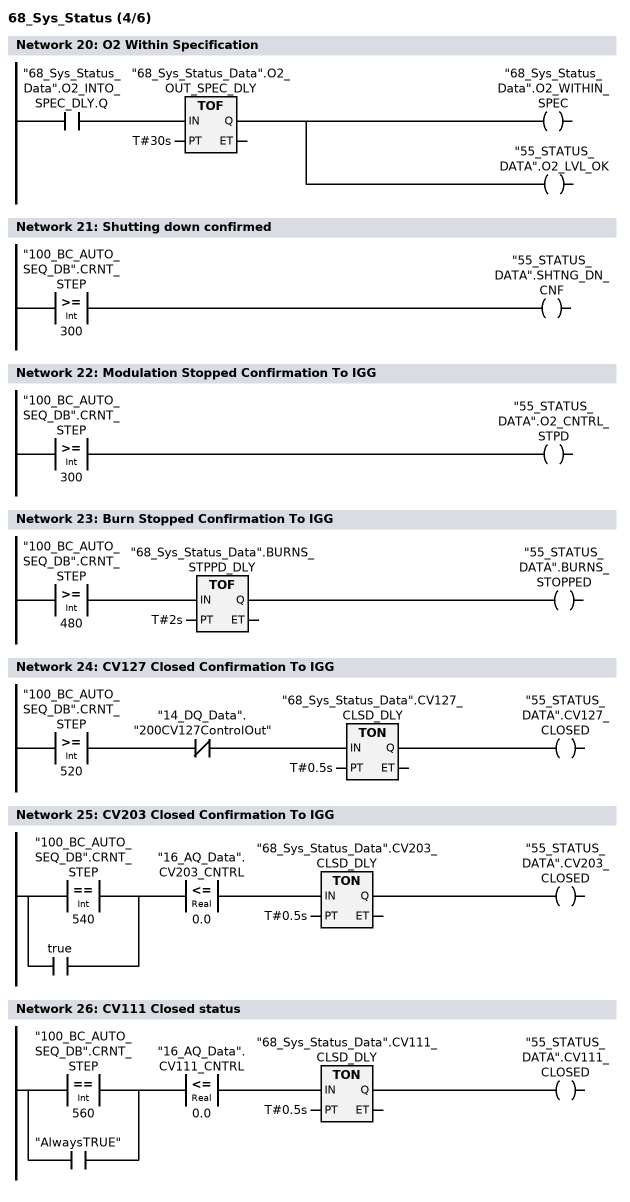
   "68_Sys_Status_Data".O2_OUT_SPEC_DLY.TOF(IN := "68_Sys_Status_Data".O2_INTO_SPEC_DLY.Q, PT := T#30s);
   "68_Sys_Status_Data".O2_WITHIN_SPEC := "68_Sys_Status_Data".O2_OUT_SPEC_DLY.Q;
   "55_STATUS_DATA".O2_LVL_OK := "68_Sys_Status_Data".O2_OUT_SPEC_DLY.Q;
END_REGION

REGION Network 21: Shutting down confirmed
   RUNG wire#powerrail
      { S7_Templates := "SrcType := Int" } GE_Contact(in1 := "100_BC_AUTO_SEQ_DB".CRNT_STEP, in2 := 300)
      Coil( "55_STATUS_DATA".SHTNG_DN_CNF )
   END_RUNG
   // the same network as SCL:
   "55_STATUS_DATA".SHTNG_DN_CNF := "100_BC_AUTO_SEQ_DB".CRNT_STEP >= 300;
END_REGION

REGION Network 22: Modulation Stopped Confirmation To IGG
   RUNG wire#powerrail
      { S7_Templates := "SrcType := Int" } GE_Contact(in1 := "100_BC_AUTO_SEQ_DB".CRNT_STEP, in2 := 300)
      Coil( "55_STATUS_DATA".O2_CNTRL_STPD )
   END_RUNG
   // the same network as SCL:
   "55_STATUS_DATA".O2_CNTRL_STPD := "100_BC_AUTO_SEQ_DB".CRNT_STEP >= 300;
END_REGION

REGION Network 23: Burn Stopped Confirmation To IGG
   "68_Sys_Status_Data".BURNS_STPPD_DLY.TOF(IN := "100_BC_AUTO_SEQ_DB".CRNT_STEP >= 480, PT := T#2s);
   "55_STATUS_DATA".BURNS_STOPPED := "68_Sys_Status_Data".BURNS_STPPD_DLY.Q;
END_REGION

REGION Network 24: CV127 Closed Confirmation To IGG
   "68_Sys_Status_Data".CV127_CLSD_DLY.TON(IN := ("100_BC_AUTO_SEQ_DB".CRNT_STEP >= 520) AND NOT "14_DQ_Data"."200CV127ControlOut",
                           PT := T#0.5s);
   "55_STATUS_DATA".CV127_CLOSED := "68_Sys_Status_Data".CV127_CLSD_DLY.Q;
END_REGION

REGION Network 25: CV203 Closed Confirmation To IGG
   "68_Sys_Status_Data".CV203_CLSD_DLY.TON(IN := (("100_BC_AUTO_SEQ_DB".CRNT_STEP = 540) OR true) AND ("16_AQ_Data".CV203_CNTRL <= 0.0),
                           PT := T#0.5s);
   "55_STATUS_DATA".CV203_CLOSED := "68_Sys_Status_Data".CV203_CLSD_DLY.Q;
END_REGION

REGION Network 26: CV111 Closed status
   "68_Sys_Status_Data".CV111_CLSD_DLY.TON(IN := (("100_BC_AUTO_SEQ_DB".CRNT_STEP = 560) OR "AlwaysTRUE") AND ("16_AQ_Data".CV111_CNTRL <= 0.0),
                           PT := T#0.5s);
   "55_STATUS_DATA".CV111_CLOSED := "68_Sys_Status_Data".CV111_CLSD_DLY.Q;
END_REGION

REGION Network 27: BC Shutdown sequence done
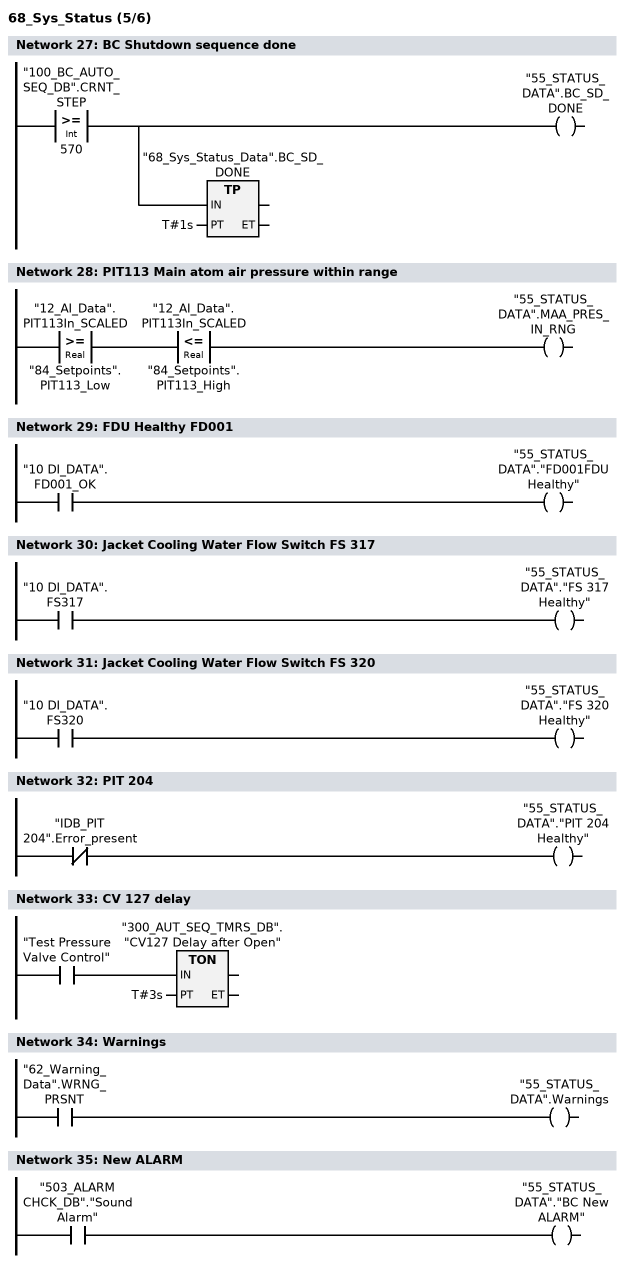
   "55_STATUS_DATA".BC_SD_DONE := "100_BC_AUTO_SEQ_DB".CRNT_STEP >= 570;
   "68_Sys_Status_Data".BC_SD_DONE.TP(IN := "55_STATUS_DATA".BC_SD_DONE, PT := T#1s);
END_REGION

REGION Network 28: PIT113 Main atom air pressure within range
   RUNG wire#powerrail
      { S7_Templates := "SrcType := Real" } GE_Contact(in1 := "12_AI_Data".PIT113In_SCALED, in2 := "84_Setpoints".PIT113_Low)
      { S7_Templates := "SrcType := Real" } LE_Contact(in1 := "12_AI_Data".PIT113In_SCALED, in2 := "84_Setpoints".PIT113_High)
      Coil( "55_STATUS_DATA".MAA_PRES_IN_RNG )
   END_RUNG
   // the same network as SCL:
   "55_STATUS_DATA".MAA_PRES_IN_RNG := ("12_AI_Data".PIT113In_SCALED >= "84_Setpoints".PIT113_Low) AND ("12_AI_Data".PIT113In_SCALED <= "84_Setpoints".PIT113_High);
END_REGION

REGION Network 29: FDU Healthy FD001
   RUNG wire#powerrail
      Contact( "10 DI_DATA".FD001_OK )
      Coil( "55_STATUS_DATA"."FD001FDU Healthy" )
   END_RUNG
   // the same network as SCL:
   "55_STATUS_DATA"."FD001FDU Healthy" := "10 DI_DATA".FD001_OK;
END_REGION

REGION Network 30: Jacket Cooling Water Flow Switch FS 317
   RUNG wire#powerrail
      Contact( "10 DI_DATA".FS317 )
      Coil( "55_STATUS_DATA"."FS 317 Healthy" )
   END_RUNG
   // the same network as SCL:
   "55_STATUS_DATA"."FS 317 Healthy" := "10 DI_DATA".FS317;
END_REGION

REGION Network 31: Jacket Cooling Water Flow Switch FS 320
   RUNG wire#powerrail
      Contact( "10 DI_DATA".FS320 )
      Coil( "55_STATUS_DATA"."FS 320 Healthy" )
   END_RUNG
   // the same network as SCL:
   "55_STATUS_DATA"."FS 320 Healthy" := "10 DI_DATA".FS320;
END_REGION

REGION Network 32: PIT 204
   RUNG wire#powerrail
      I_Contact( "IDB_PIT 204".Error_present )
      Coil( "55_STATUS_DATA"."PIT 204 Healthy" )
   END_RUNG
   // the same network as SCL:
   "55_STATUS_DATA"."PIT 204 Healthy" := NOT "IDB_PIT 204".Error_present;
END_REGION

REGION Network 33: CV 127 delay
   "300_AUT_SEQ_TMRS_DB"."CV127 Delay after Open".TON(IN := "Test Pressure Valve Control", PT := T#3s);
END_REGION

REGION Network 34: Warnings
   RUNG wire#powerrail
      Contact( "62_Warning_Data".WRNG_PRSNT )
      Coil( "55_STATUS_DATA".Warnings )
   END_RUNG
   // the same network as SCL:
   "55_STATUS_DATA".Warnings := "62_Warning_Data".WRNG_PRSNT;
END_REGION

REGION Network 35: New ALARM
   RUNG wire#powerrail
      Contact( "503_ALARM CHCK_DB"."Sound Alarm" )
      Coil( "55_STATUS_DATA"."BC New ALARM" )
   END_RUNG
   // the same network as SCL:
   "55_STATUS_DATA"."BC New ALARM" := "503_ALARM CHCK_DB"."Sound Alarm";
END_REGION

REGION Network 36: New WARNING
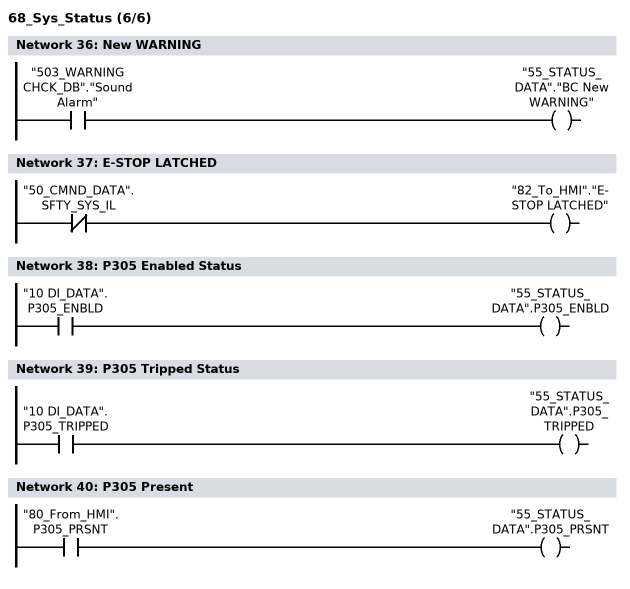
   RUNG wire#powerrail
      Contact( "503_WARNING CHCK_DB"."Sound Alarm" )
      Coil( "55_STATUS_DATA"."BC New WARNING" )
   END_RUNG
   // the same network as SCL:
   "55_STATUS_DATA"."BC New WARNING" := "503_WARNING CHCK_DB"."Sound Alarm";
END_REGION

REGION Network 37: E-STOP LATCHED
   RUNG wire#powerrail
      I_Contact( "50_CMND_DATA".SFTY_SYS_IL )
      Coil( "82_To_HMI"."E-STOP LATCHED" )
   END_RUNG
   // the same network as SCL:
   "82_To_HMI"."E-STOP LATCHED" := NOT "50_CMND_DATA".SFTY_SYS_IL;
END_REGION

REGION Network 38: P305 Enabled Status
   RUNG wire#powerrail
      Contact( "10 DI_DATA".P305_ENBLD )
      Coil( "55_STATUS_DATA".P305_ENBLD )
   END_RUNG
   // the same network as SCL:
   "55_STATUS_DATA".P305_ENBLD := "10 DI_DATA".P305_ENBLD;
END_REGION

REGION Network 39: P305 Tripped Status
   RUNG wire#powerrail
      Contact( "10 DI_DATA".P305_TRIPPED )
      Coil( "55_STATUS_DATA".P305_TRIPPED )
   END_RUNG
   // the same network as SCL:
   "55_STATUS_DATA".P305_TRIPPED := "10 DI_DATA".P305_TRIPPED;
END_REGION

REGION Network 40: P305 Present
   RUNG wire#powerrail
      Contact( "80_From_HMI".P305_PRSNT )
      Coil( "55_STATUS_DATA".P305_PRSNT )
   END_RUNG
   // the same network as SCL:
   "55_STATUS_DATA".P305_PRSNT := "80_From_HMI".P305_PRSNT;
END_REGION
END_FUNCTION

// folder: 70 - 79 Modes of Operation

FUNCTION "70_Mode_Control" : Void   // FC70, LAD
TITLE = Mode Control
{ S7_Optimized_Access := 'TRUE' }
AUTHOR : JRS
VERSION : 0.1
// To determine the current mode of operation 1=Auto(default), 2=Manual, 3=FatAuto, 4=FatManual
   VAR_TEMP   // added for the SCL form of the ladder/FBD networks
      _w1 : Bool;
   END_VAR
BEGIN

REGION Network 1: Default = Automatic
   // Set default to Automatic (on first scan)
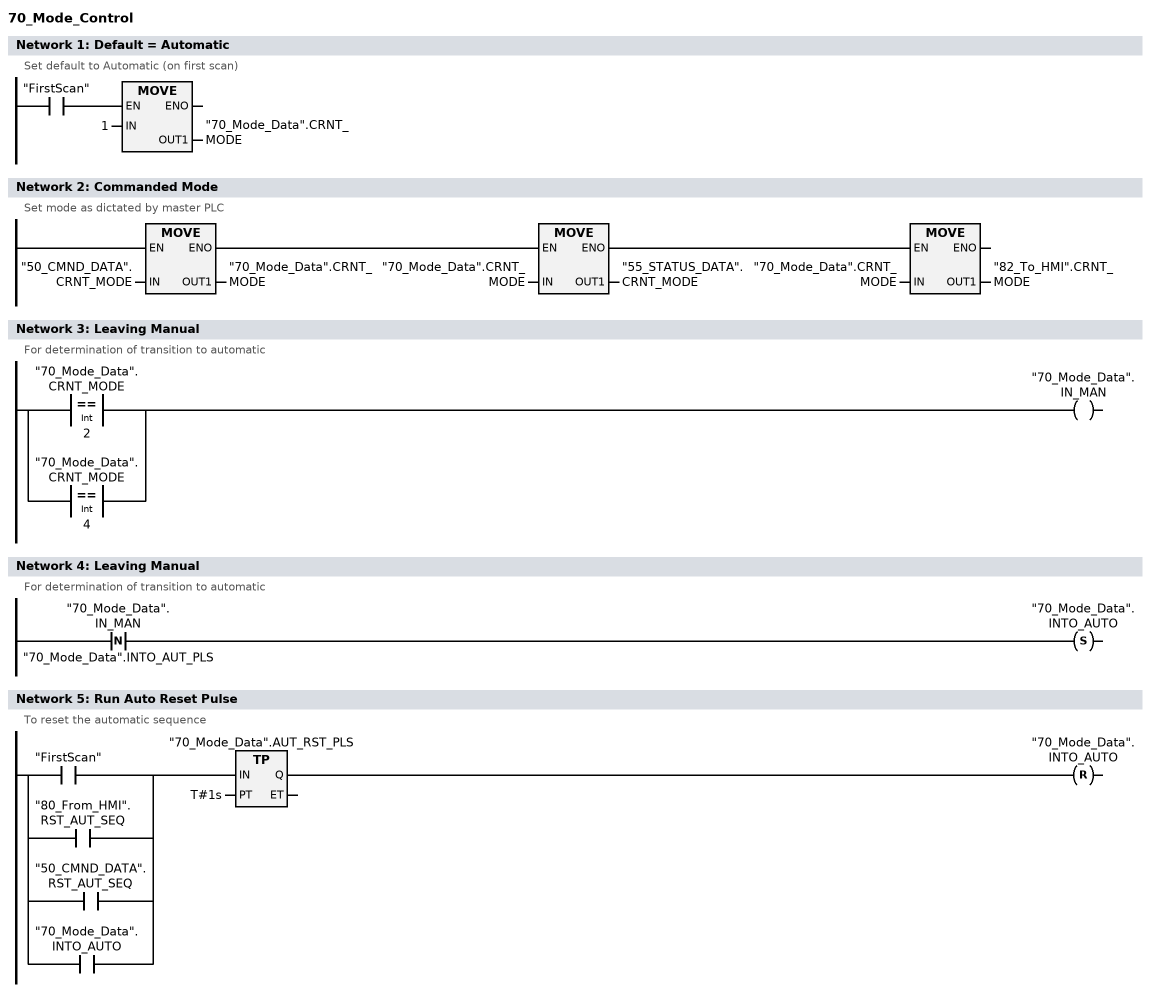
   RUNG wire#powerrail
      Contact( "FirstScan" )
      Move(in := 1, out1 => "70_Mode_Data".CRNT_MODE)
   END_RUNG
   // the same network as SCL:
   IF "FirstScan" THEN "70_Mode_Data".CRNT_MODE := 1; END_IF;
END_REGION

REGION Network 2: Commanded Mode
   // Set mode as dictated by master PLC
   RUNG wire#powerrail
      Move(in := "50_CMND_DATA".CRNT_MODE, out1 => "70_Mode_Data".CRNT_MODE)
      Move(in := "70_Mode_Data".CRNT_MODE, out1 => "55_STATUS_DATA".CRNT_MODE)
      Move(in := "70_Mode_Data".CRNT_MODE, out1 => "82_To_HMI".CRNT_MODE)
   END_RUNG
   // the same network as SCL:
   "70_Mode_Data".CRNT_MODE := "50_CMND_DATA".CRNT_MODE;
   "55_STATUS_DATA".CRNT_MODE := "70_Mode_Data".CRNT_MODE;
   "82_To_HMI".CRNT_MODE := "70_Mode_Data".CRNT_MODE;
END_REGION

REGION Network 3: Leaving Manual
   // For determination of transition to automatic
   RUNG wire#powerrail
      { S7_Templates := "SrcType := Int" } EQ_Contact(in1 := "70_Mode_Data".CRNT_MODE, in2 := 2)
      wire#w1
      Coil( "70_Mode_Data".IN_MAN )
   END_RUNG
   RUNG wire#powerrail
      { S7_Templates := "SrcType := Int" } EQ_Contact(in1 := "70_Mode_Data".CRNT_MODE, in2 := 4)
   END_RUNG wire#w1
   // the same network as SCL:
   "70_Mode_Data".IN_MAN := ("70_Mode_Data".CRNT_MODE = 2) OR ("70_Mode_Data".CRNT_MODE = 4);
END_REGION

REGION Network 4: Leaving Manual
   // For determination of transition to automatic
   RUNG wire#powerrail
      N_Contact(operand := "70_Mode_Data".IN_MAN, bit := "70_Mode_Data".INTO_AUT_PLS)
      S_Coil( "70_Mode_Data".INTO_AUTO )
   END_RUNG
   // the same network as SCL:
   #_w1 := NOT "70_Mode_Data".IN_MAN AND "70_Mode_Data".INTO_AUT_PLS;   // falling edge of "70_Mode_Data".IN_MAN
   "70_Mode_Data".INTO_AUT_PLS := "70_Mode_Data".IN_MAN;
   IF #_w1 THEN "70_Mode_Data".INTO_AUTO := TRUE; END_IF;
END_REGION

REGION Network 5: Run Auto Reset Pulse
   // To reset the automatic sequence
   "70_Mode_Data".AUT_RST_PLS.TP(IN := "FirstScan" OR "80_From_HMI".RST_AUT_SEQ OR "50_CMND_DATA".RST_AUT_SEQ OR "70_Mode_Data".INTO_AUTO,
                           PT := T#1s);
   IF "70_Mode_Data".AUT_RST_PLS.Q THEN "70_Mode_Data".INTO_AUTO := FALSE; END_IF;
END_REGION
END_FUNCTION

// folder: 90 - 99 Manual Functions

FUNCTION "90_Manual_Control" : Void   // FC90, LAD
TITLE = Manual Control
{ S7_Optimized_Access := 'TRUE' }
AUTHOR : JHT
VERSION : 0.1
// Code for manual operation of equipment
   VAR_TEMP   // added for the SCL form of the ladder/FBD networks
      _w1 : Bool;
      _w2 : Bool;
      _w3 : Bool;
      _w4 : Bool;
      _w5 : Bool;
      _w6 : Bool;
   END_VAR
BEGIN

REGION Network 1: Zero Auto Step Numbers
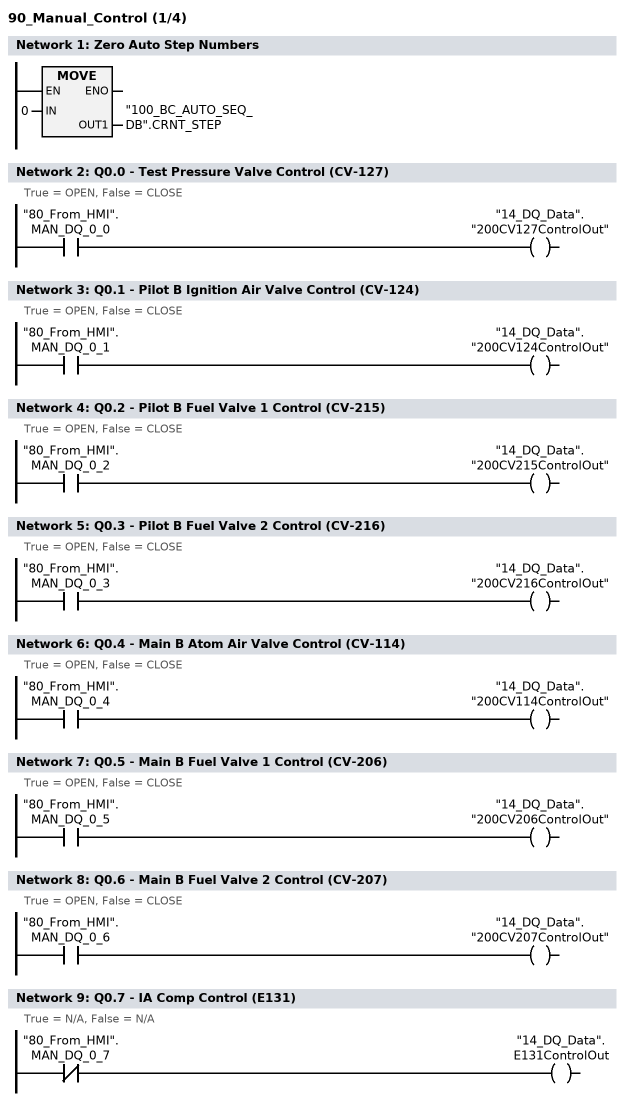
   RUNG wire#powerrail
      Move(in := 0, out1 => "100_BC_AUTO_SEQ_DB".CRNT_STEP)
   END_RUNG
   // the same network as SCL:
   "100_BC_AUTO_SEQ_DB".CRNT_STEP := 0;
END_REGION

REGION Network 2: Q0.0 - Test Pressure Valve Control (CV-127)
   // True = OPEN, False = CLOSE
   RUNG wire#powerrail
      Contact( "80_From_HMI".MAN_DQ_0_0 )
      Coil( "14_DQ_Data"."200CV127ControlOut" )
   END_RUNG
   // the same network as SCL:
   "14_DQ_Data"."200CV127ControlOut" := "80_From_HMI".MAN_DQ_0_0;
END_REGION

REGION Network 3: Q0.1 - Pilot B Ignition Air Valve Control (CV-124)
   // True = OPEN, False = CLOSE
   RUNG wire#powerrail
      Contact( "80_From_HMI".MAN_DQ_0_1 )
      Coil( "14_DQ_Data"."200CV124ControlOut" )
   END_RUNG
   // the same network as SCL:
   "14_DQ_Data"."200CV124ControlOut" := "80_From_HMI".MAN_DQ_0_1;
END_REGION

REGION Network 4: Q0.2 - Pilot B Fuel Valve 1 Control (CV-215)
   // True = OPEN, False = CLOSE
   RUNG wire#powerrail
      Contact( "80_From_HMI".MAN_DQ_0_2 )
      Coil( "14_DQ_Data"."200CV215ControlOut" )
   END_RUNG
   // the same network as SCL:
   "14_DQ_Data"."200CV215ControlOut" := "80_From_HMI".MAN_DQ_0_2;
END_REGION

REGION Network 5: Q0.3 - Pilot B Fuel Valve 2 Control (CV-216)
   // True = OPEN, False = CLOSE
   RUNG wire#powerrail
      Contact( "80_From_HMI".MAN_DQ_0_3 )
      Coil( "14_DQ_Data"."200CV216ControlOut" )
   END_RUNG
   // the same network as SCL:
   "14_DQ_Data"."200CV216ControlOut" := "80_From_HMI".MAN_DQ_0_3;
END_REGION

REGION Network 6: Q0.4 - Main B Atom Air Valve Control (CV-114)
   // True = OPEN, False = CLOSE
   RUNG wire#powerrail
      Contact( "80_From_HMI".MAN_DQ_0_4 )
      Coil( "14_DQ_Data"."200CV114ControlOut" )
   END_RUNG
   // the same network as SCL:
   "14_DQ_Data"."200CV114ControlOut" := "80_From_HMI".MAN_DQ_0_4;
END_REGION

REGION Network 7: Q0.5 - Main B Fuel Valve 1 Control (CV-206)
   // True = OPEN, False = CLOSE
   RUNG wire#powerrail
      Contact( "80_From_HMI".MAN_DQ_0_5 )
      Coil( "14_DQ_Data"."200CV206ControlOut" )
   END_RUNG
   // the same network as SCL:
   "14_DQ_Data"."200CV206ControlOut" := "80_From_HMI".MAN_DQ_0_5;
END_REGION

REGION Network 8: Q0.6 - Main B Fuel Valve 2 Control (CV-207)
   // True = OPEN, False = CLOSE
   RUNG wire#powerrail
      Contact( "80_From_HMI".MAN_DQ_0_6 )
      Coil( "14_DQ_Data"."200CV207ControlOut" )
   END_RUNG
   // the same network as SCL:
   "14_DQ_Data"."200CV207ControlOut" := "80_From_HMI".MAN_DQ_0_6;
END_REGION

REGION Network 9: Q0.7 - IA Comp Control (E131)
   // True = N/A, False = N/A
   RUNG wire#powerrail
      I_Contact( "80_From_HMI".MAN_DQ_0_7 )
      Coil( "14_DQ_Data".E131ControlOut )
   END_RUNG
   // the same network as SCL:
   "14_DQ_Data".E131ControlOut := NOT "80_From_HMI".MAN_DQ_0_7;
END_REGION

REGION Network 10: Q1.0 - CSW Pump Control (P301)
   // True = N/A, False = N/A
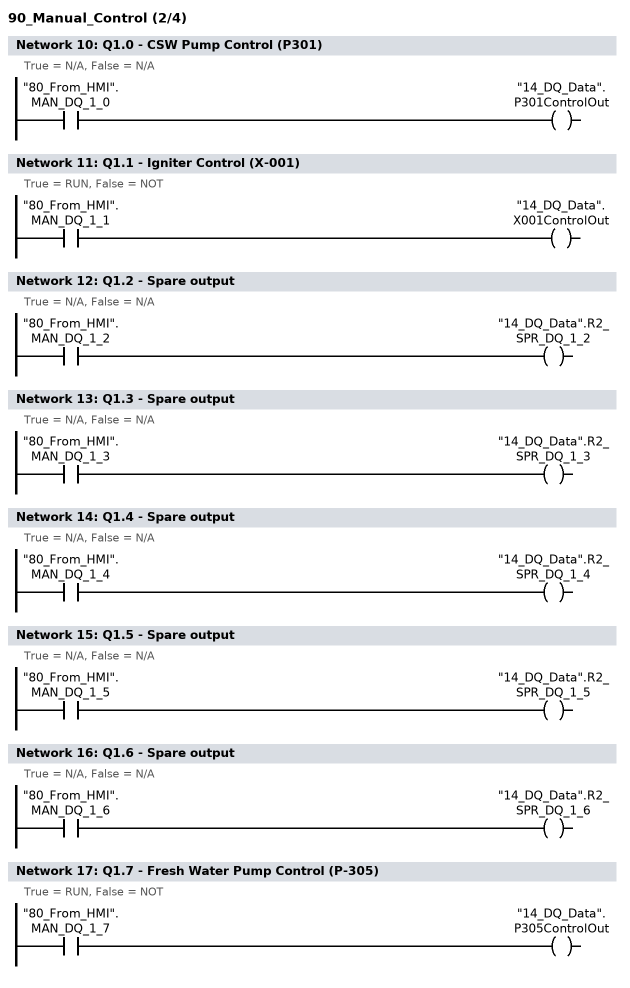
   RUNG wire#powerrail
      Contact( "80_From_HMI".MAN_DQ_1_0 )
      Coil( "14_DQ_Data".P301ControlOut )
   END_RUNG
   // the same network as SCL:
   "14_DQ_Data".P301ControlOut := "80_From_HMI".MAN_DQ_1_0;
END_REGION

REGION Network 11: Q1.1 - Igniter Control (X-001)
   // True = RUN, False = NOT
   RUNG wire#powerrail
      Contact( "80_From_HMI".MAN_DQ_1_1 )
      Coil( "14_DQ_Data".X001ControlOut )
   END_RUNG
   // the same network as SCL:
   "14_DQ_Data".X001ControlOut := "80_From_HMI".MAN_DQ_1_1;
END_REGION

REGION Network 12: Q1.2 - Spare output
   // True = N/A, False = N/A
   RUNG wire#powerrail
      Contact( "80_From_HMI".MAN_DQ_1_2 )
      Coil( "14_DQ_Data".R2_SPR_DQ_1_2 )
   END_RUNG
   // the same network as SCL:
   "14_DQ_Data".R2_SPR_DQ_1_2 := "80_From_HMI".MAN_DQ_1_2;
END_REGION

REGION Network 13: Q1.3 - Spare output
   // True = N/A, False = N/A
   RUNG wire#powerrail
      Contact( "80_From_HMI".MAN_DQ_1_3 )
      Coil( "14_DQ_Data".R2_SPR_DQ_1_3 )
   END_RUNG
   // the same network as SCL:
   "14_DQ_Data".R2_SPR_DQ_1_3 := "80_From_HMI".MAN_DQ_1_3;
END_REGION

REGION Network 14: Q1.4 - Spare output
   // True = N/A, False = N/A
   RUNG wire#powerrail
      Contact( "80_From_HMI".MAN_DQ_1_4 )
      Coil( "14_DQ_Data".R2_SPR_DQ_1_4 )
   END_RUNG
   // the same network as SCL:
   "14_DQ_Data".R2_SPR_DQ_1_4 := "80_From_HMI".MAN_DQ_1_4;
END_REGION

REGION Network 15: Q1.5 - Spare output
   // True = N/A, False = N/A
   RUNG wire#powerrail
      Contact( "80_From_HMI".MAN_DQ_1_5 )
      Coil( "14_DQ_Data".R2_SPR_DQ_1_5 )
   END_RUNG
   // the same network as SCL:
   "14_DQ_Data".R2_SPR_DQ_1_5 := "80_From_HMI".MAN_DQ_1_5;
END_REGION

REGION Network 16: Q1.6 - Spare output
   // True = N/A, False = N/A
   RUNG wire#powerrail
      Contact( "80_From_HMI".MAN_DQ_1_6 )
      Coil( "14_DQ_Data".R2_SPR_DQ_1_6 )
   END_RUNG
   // the same network as SCL:
   "14_DQ_Data".R2_SPR_DQ_1_6 := "80_From_HMI".MAN_DQ_1_6;
END_REGION

REGION Network 17: Q1.7 - Fresh Water Pump Control (P-305)
   // True = RUN, False = NOT
   RUNG wire#powerrail
      Contact( "80_From_HMI".MAN_DQ_1_7 )
      Coil( "14_DQ_Data".P305ControlOut )
   END_RUNG
   // the same network as SCL:
   "14_DQ_Data".P305ControlOut := "80_From_HMI".MAN_DQ_1_7;
END_REGION

REGION Network 18: QW96 - Spare Output (Hardware Channel De-activated)
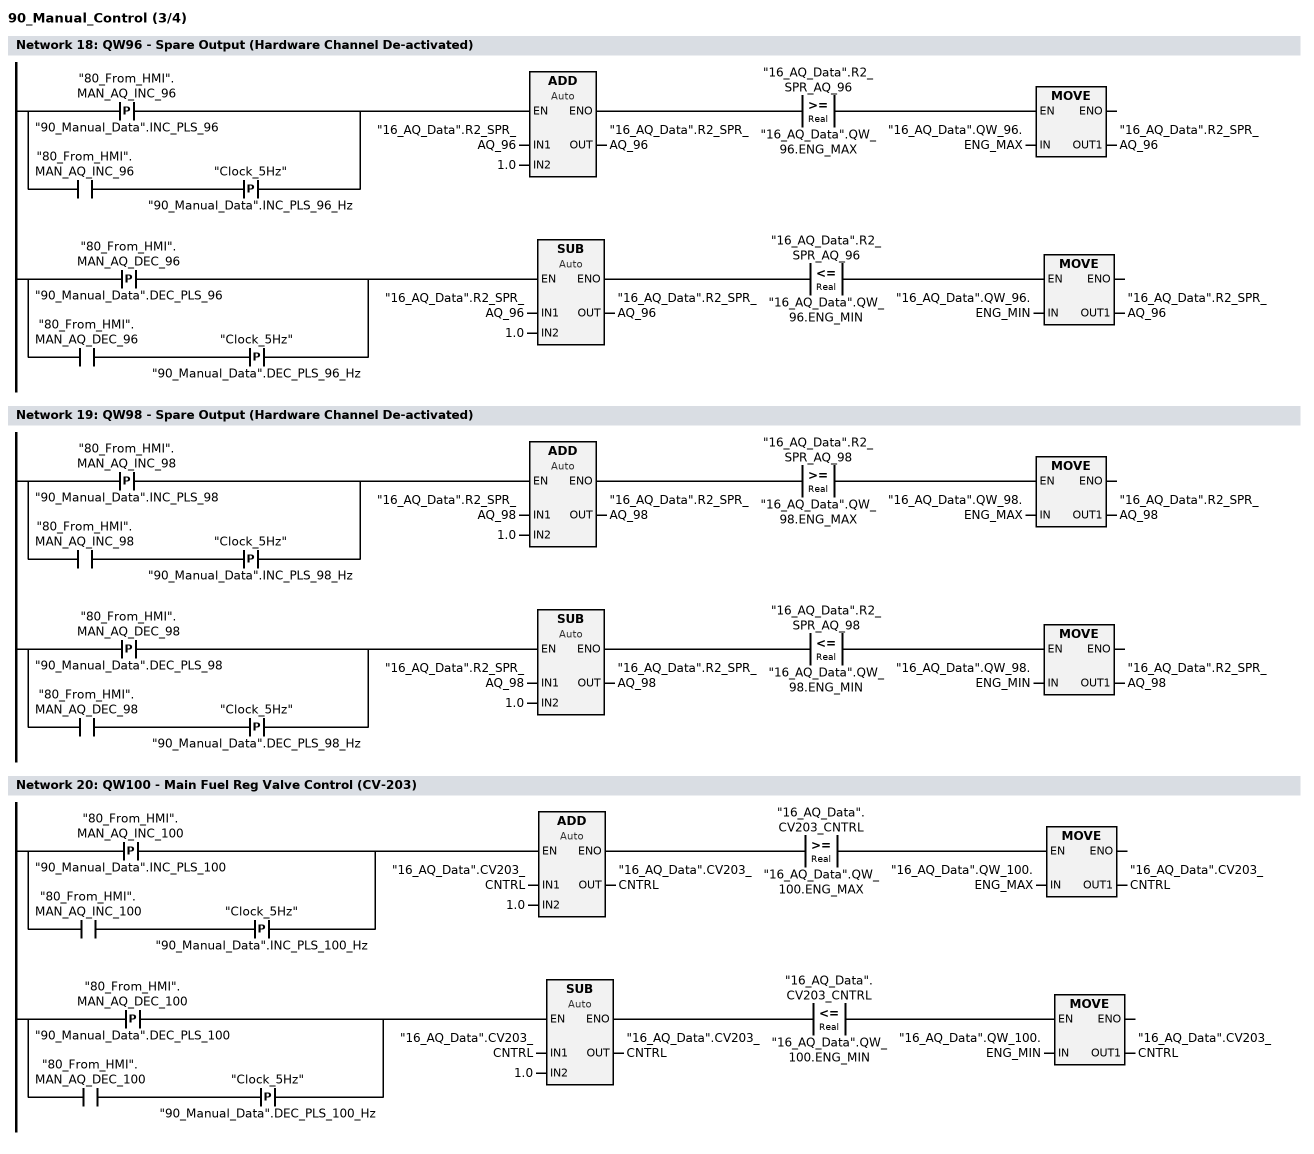
   RUNG wire#powerrail
      P_Contact(operand := "80_From_HMI".MAN_AQ_INC_96, bit := "90_Manual_Data".INC_PLS_96)
      wire#w1
      Add(in1 := "16_AQ_Data".R2_SPR_AQ_96, in2 := 1.0, out => "16_AQ_Data".R2_SPR_AQ_96)
      { S7_Templates := "SrcType := Real" } GE_Contact(in1 := "16_AQ_Data".R2_SPR_AQ_96, in2 := "16_AQ_Data".QW_96.ENG_MAX)
      { S7_GenerateENO := "TRUE" } Move(in := "16_AQ_Data".QW_96.ENG_MAX, out1 => "16_AQ_Data".R2_SPR_AQ_96)
   END_RUNG
   RUNG wire#powerrail
      Contact( "80_From_HMI".MAN_AQ_INC_96 )
      P_Contact(operand := "Clock_5Hz", bit := "90_Manual_Data".INC_PLS_96_Hz)
   END_RUNG wire#w1
   RUNG wire#powerrail
      P_Contact(operand := "80_From_HMI".MAN_AQ_DEC_96, bit := "90_Manual_Data".DEC_PLS_96)
      wire#w2
      Sub(in1 := "16_AQ_Data".R2_SPR_AQ_96, in2 := 1.0, out => "16_AQ_Data".R2_SPR_AQ_96)
      { S7_Templates := "SrcType := Real" } LE_Contact(in1 := "16_AQ_Data".R2_SPR_AQ_96, in2 := "16_AQ_Data".QW_96.ENG_MIN)
      { S7_GenerateENO := "TRUE" } Move(in := "16_AQ_Data".QW_96.ENG_MIN, out1 => "16_AQ_Data".R2_SPR_AQ_96)
   END_RUNG
   RUNG wire#powerrail
      Contact( "80_From_HMI".MAN_AQ_DEC_96 )
      P_Contact(operand := "Clock_5Hz", bit := "90_Manual_Data".DEC_PLS_96_Hz)
   END_RUNG wire#w2
   // the same network as SCL:
   #_w1 := "80_From_HMI".MAN_AQ_INC_96 AND NOT "90_Manual_Data".INC_PLS_96;   // rising edge of "80_From_HMI".MAN_AQ_INC_96
   "90_Manual_Data".INC_PLS_96 := "80_From_HMI".MAN_AQ_INC_96;
   #_w2 := "80_From_HMI".MAN_AQ_INC_96 AND "Clock_5Hz" AND NOT "90_Manual_Data".INC_PLS_96_Hz;   // rising edge of "Clock_5Hz"
   "90_Manual_Data".INC_PLS_96_Hz := "Clock_5Hz";
   #_w3 := #_w1 OR #_w2;
   IF #_w3 THEN "16_AQ_Data".R2_SPR_AQ_96 := "16_AQ_Data".R2_SPR_AQ_96 + 1.0; END_IF;
   IF #_w3 AND ("16_AQ_Data".R2_SPR_AQ_96 >= "16_AQ_Data".QW_96.ENG_MAX) THEN
       "16_AQ_Data".R2_SPR_AQ_96 := "16_AQ_Data".QW_96.ENG_MAX;
   END_IF;
   #_w4 := "80_From_HMI".MAN_AQ_DEC_96 AND NOT "90_Manual_Data".DEC_PLS_96;   // rising edge of "80_From_HMI".MAN_AQ_DEC_96
   "90_Manual_Data".DEC_PLS_96 := "80_From_HMI".MAN_AQ_DEC_96;
   #_w5 := "80_From_HMI".MAN_AQ_DEC_96 AND "Clock_5Hz" AND NOT "90_Manual_Data".DEC_PLS_96_Hz;   // rising edge of "Clock_5Hz"
   "90_Manual_Data".DEC_PLS_96_Hz := "Clock_5Hz";
   #_w6 := #_w4 OR #_w5;
   IF #_w6 THEN "16_AQ_Data".R2_SPR_AQ_96 := "16_AQ_Data".R2_SPR_AQ_96 - 1.0; END_IF;
   IF #_w6 AND ("16_AQ_Data".R2_SPR_AQ_96 <= "16_AQ_Data".QW_96.ENG_MIN) THEN
       "16_AQ_Data".R2_SPR_AQ_96 := "16_AQ_Data".QW_96.ENG_MIN;
   END_IF;
END_REGION
